   hm 20. oct. 2006 rev 1.5
    changed time_zone_offset from Real to INT, now in Minutes

   hm 27. feb. 2009 rev 1.6
    added type conversions to avoid warnings under codesys 3.0

   ks 13. nov. 2009 rev 1.7
    corrected error in formula

   *)
END_FUNCTION

FUNCTION "MINUTE" : Int   // FC197, SCL
TITLE = MINUTE
{ S7_Optimized_Access := 'FALSE' }
AUTHOR : hugo
FAMILY : TIDT
NAME : MINUTE
VERSION : 1.1
// extracts the minutes out of TOD truncating the ceconds
   VAR_INPUT
      itod : Time_Of_Day;
   END_VAR
BEGIN


     #MINUTE := DINT_TO_INT(T_CONV(#itod)/60000 - T_CONV(#itod)/3600000 * 60);


   (* change history

   2.10.2006 changes name of input to itod

   *)
END_FUNCTION

FUNCTION "MINUTE_OF_DT" : Int   // FC198, SCL
TITLE = MINUTE_OF_DT
{ S7_Optimized_Access := 'FALSE' }
AUTHOR : oscat
FAMILY : TIDT
NAME : M_DT
VERSION : 1.0
// MINUTE_OF_DT returns the current minute (minute of the hour) of a DT variable
   VAR_INPUT
      XDT : Date_And_Time;
      _XDT AT XDT : Array[0..7] of Byte;
   END_VAR
BEGIN


   #MINUTE_OF_DT := BCD16_TO_INT(#_XDT[4]); 

   (*
       original code:
       MINUTE_OF_DT := DWORD_TO_INT(DT_TO_DWORD(XDT) MOD 3600)/60;
   *)

   (* revision history
   hm      6.9.2008    rev 1.0
       original version


   *)
END_FUNCTION

FUNCTION "MINUTE_TO_TIME" : Time   // FC199, SCL
TITLE = MINUTE_TO_TIME
{ S7_Optimized_Access := 'FALSE' }
AUTHOR : hugo
FAMILY : TIDT
NAME : MIN2TI
VERSION : 1.2
// converts an amount of minutes in real to time
   VAR_INPUT
      IN : Real;
   END_VAR
BEGIN


   #MINUTE_TO_TIME := T_CONV(REAL_TO_DINT(#IN * 60000));


   (* revision history
   hm  4. aug 2006 rev 1.0
       original version

   hm  14. mar 2008    rev 1.1
       rounded the input after the last digit

   hm  24. feb. 2009   rev 1.2
       changed input to IN

   *)
END_FUNCTION

FUNCTION "MONTH_BEGIN" : Date   // FC200, SCL
TITLE = MONTH_BEGIN
{ S7_Optimized_Access := 'FALSE' }
AUTHOR : hugo
FAMILY : TIDT
NAME : MONBEG
VERSION : 1.0
// returns the date for the first day of the current month in the current year.
// 
// uses: DINT_DATE [FC404]
//       DATE_DINT [FC405]
//       DAY_OF_MONTH [FC178]
//       DAY_OF_YEAR [FC180] 
//       YEAR_BEGIN [FC217]
//       YEAR_OF_DATE [FC219]
//       LEAP_OF_DATE [FC193] 
//       LEAP_YEAR [FC194]
   VAR_INPUT
      idate : Date;
   END_VAR
BEGIN


   #MONTH_BEGIN := "DINT_DATE"("DATE_DINT"(#idate) - ("DAY_OF_MONTH"(#idate) - 1) * 86400);



   (* revision history
   hm  15. JUN: 2008   rev 1.0
       original version 


   *)
END_FUNCTION

FUNCTION "MONTH_END" : Date   // FC201, SCL
TITLE = MONTH_END
{ S7_Optimized_Access := 'FALSE' }
AUTHOR : hugo
FAMILY : TIDT
NAME : MONEND
VERSION : 1.1
// returns the date for the first day of the current month in the current year.
// 
// uses: DINT_DATE [FC404]
//       DATE_DINT [FC405]
//       SET_DATE [FC213]
//       LEAP_YEAR [FC194] 
//       YEAR_OF_DATE [FC219]
//       MONTH_OF_DATE [FC202]
//       DAY_OF_YEAR [FC180] 
//       YEAR_BEGIN [FC217]
//       LEAP_OF_DATE [FC193]
   VAR_INPUT
      idate : Date;
   END_VAR
BEGIN


   #MONTH_END := "DINT_DATE"("DATE_DINT"("SET_DATE"(YEAR:="YEAR_OF_DATE"(#idate),MONTH:="MONTH_OF_DATE"(#idate)+1,DAY:=1)) - 86400);

   (* revision history
   hm  15. jun. 2008   rev 1.0
       original version    

   hm  7. oct. 2008    rev 1.1
       changed function year to year_of_date
       changed function month to month_of_date

   *)
END_FUNCTION

FUNCTION "MONTH_OF_DATE" : Int   // FC202, SCL
TITLE = MONTH_OF_DATE
{ S7_Optimized_Access := 'FALSE' }
AUTHOR : hugo
FAMILY : TIDT
NAME : MONTH
VERSION : 1.3
// returns the month of a date  
// 
// uses: DAY_OF_YEAR [FC180]
//       YEAR_BEGIN [FC217] 
//       YEAR_OF_DATE [FC219] 
//       LEAP_OF_DATE [FC193]
//       LEAP_YEAR [FC194]
   VAR_INPUT
      IDATE : Date;
   END_VAR
BEGIN


   #MONTH_OF_DATE := "DAY_OF_YEAR"(#IDATE);
   IF #MONTH_OF_DATE < 32 THEN
       #MONTH_OF_DATE := 1;
   ELSIF "LEAP_OF_DATE"(#IDATE) THEN
       #MONTH_OF_DATE := (#MONTH_OF_DATE * 53 + 1668) / 1623;
   ELSE
       #MONTH_OF_DATE := (#MONTH_OF_DATE * 53 + 1700) / 1620;
   END_IF;


   (* code for rev 1.2
   MONTH_OF_DATE := DAY_OF_YEAR(IDATE);
   IF LEAP_OF_DATE(IDATE) THEN
       CASE MONTH_OF_DATE OF
           1..31   :   MONTH_OF_DATE := 1;
           32..60  :   MONTH_OF_DATE := 2;
           61..91  :   MONTH_OF_DATE := 3;
           92..121 :   MONTH_OF_DATE := 4;
           122..152:   MONTH_OF_DATE := 5;
           153..182:   MONTH_OF_DATE := 6;
           183..213:   MONTH_OF_DATE := 7;
           214..244:   MONTH_OF_DATE := 8;
           245..274:   MONTH_OF_DATE := 9;
           275..305:   MONTH_OF_DATE := 10;
           306..335:   MONTH_OF_DATE := 11;
           336..366:   MONTH_OF_DATE := 12;
       END_CASE;
   ELSE
       CASE MONTH_OF_DATE OF
           1..31   :   MONTH_OF_DATE := 1;
           32..59  :   MONTH_OF_DATE := 2;
           60..90  :   MONTH_OF_DATE := 3;
           91..120 :   MONTH_OF_DATE := 4;
           121..151:   MONTH_OF_DATE := 5;
           152..181:   MONTH_OF_DATE := 6;
           182..212:   MONTH_OF_DATE := 7;
           213..243:   MONTH_OF_DATE := 8;
           244..273:   MONTH_OF_DATE := 9;
           274..304:   MONTH_OF_DATE := 10;
           305..334:   MONTH_OF_DATE := 11;
           335..365:   MONTH_OF_DATE := 12;
       END_CASE;
   END_IF;
   *)


   (* revision history
   hm  1. aug 2006 rev 1.0
       original version    

   hm  1. okt 2007 rev 1.1
       replaced old code (string conversion) with mathematics
       the execution time is now multiple times faster.

   hm  7. oct. 2008    rev 1.2
       changed name of function from month to MONTH_OF_DATE

   hm  27. mar. 2009   rev 1.3
       new improved code

   *)
END_FUNCTION

FUNCTION "MULTIME" : Time   // FC203, SCL
TITLE = MULTIME
{ S7_Optimized_Access := 'FALSE' }
AUTHOR : hugo
FAMILY : TIDT
NAME : MULTIME
VERSION : 1.1
// multiplies a time by a real number and returns a time
   VAR_INPUT
      t : Time;
      "M" : Real;
   END_VAR
BEGIN


     #MULTIME := T_CONV(REAL_TO_DINT(DINT_TO_REAL(T_CONV(#t)) * #"M"));

   (* revision history
   hm      2. oct 2006 rev 1.0
       original version

   hm      14. mar 2008    rev 1.1
       rounded the result after the last digit

   *)
END_FUNCTION

FUNCTION "PERIOD" : Bool   // FC204, SCL
TITLE = PERIOD
{ S7_Optimized_Access := 'FALSE' }
AUTHOR : hugo
FAMILY : TIDT
NAME : PERIOD
VERSION : 1.3
// PERIOD checks if a given date is between two dates (d1 and d2) d1 is the starting date and d2 the last date for the period.
// the years of the dates are ignored, so the function period cheks for a time period within a year independet of the year.
// 
// uses: DAY_OF_YEAR [FC180]
//       YEAR_BEGIN [FC217] 
//       YEAR_OF_DATE [FC219] 
//       LEAP_OF_DATE [FC193]
//       LEAP_YEAR [FC194]
   VAR_INPUT
      d1 : Date;
      dx : Date;
      d2 : Date;
   END_VAR
   VAR_TEMP
      day1 : Int;
      day2 : Int;
      dayx : Int;
   END_VAR
BEGIN


   #day1 := "DAY_OF_YEAR"(#d1);
   #day2 := "DAY_OF_YEAR"(#d2);
   #dayx := "DAY_OF_YEAR"(#dx);
   IF NOT "LEAP_OF_DATE"(#dx) AND #dayx > 58 THEN #dayx := #dayx + 1; END_IF;
   IF NOT "LEAP_OF_DATE"(#d1) AND #day1 > 58 THEN #day1 := #day1 + 1; END_IF;
   IF NOT "LEAP_OF_DATE"(#d2) AND #day2 > 58 THEN #day2 := #day2 + 1; END_IF;

   IF #day2 < #day1 THEN
       (* the period spans over the new year *)
       #PERIOD := #dayx <= #day2 OR #dayx >= #day1;
   ELSE
       #PERIOD := #dayx >= #day1 AND #dayx <= #day2;
   END_IF;

   (* code before rev 1.2
   yx := year(dx);
   p1 := date_add(d1,0,0,0,yx - year(d1));
   p2 := date_add(d2,0,0,0,yx - year(d2));

   IF p2 >= p1 THEN
       period := dx <= p2  AND dx >= p1;
   ELSE
       period := dx <= p2 OR dx >= p1;
   END_IF;
   *)


   (* revision history

   hm      19. sep 2007    rev 1.0
       original version

   hm      20. sep 2007    rev 1.1
       corrected a problem with leap year

   hm      4. jan 2008     rev 1.2
       changed code for better performance

   hm      22. mar. 2008   rev 1.3
       function would deliver wrong results when d1, d2 or dx are a leap_year

   *)
END_FUNCTION

FUNCTION "PERIOD2" : Bool   // FC205, SCL
TITLE = PERIOD2
{ S7_Optimized_Access := 'FALSE' }
AUTHOR : hugo
FAMILY : TIDT
NAME : PERIOD2
VERSION : 1.0
// PERIOD2 checks if DX is within one of 4 periods and sets the output true if so.
   VAR_INPUT
      DP : Array[0..3, 0..1] of Date;
      DX : Date;
   END_VAR
BEGIN


   #PERIOD2 :=  (#DX >= #DP[0,0] AND #DX <= #DP[0,1]) OR
               (#DX >= #DP[1,0] AND #DX <= #DP[1,1]) OR
               (#DX >= #DP[2,0] AND #DX <= #DP[2,1]) OR
               (#DX >= #DP[3,0] AND #DX <= #DP[3,1]);


   (* revision history

   hm      27. apr 2008    rev 1.0
       original version


   *)
END_FUNCTION

FUNCTION "REFRACTION" : Real   // FC206, SCL
TITLE = REFRACTION
{ S7_Optimized_Access := 'FALSE' }
AUTHOR : hugo
FAMILY : TIDT
NAME : REFRACT
VERSION : 1.1
// REFRACTION calculates the atmospheric refraction in degrees.
// the input nangle goes from 0 at the hirizon to 90 at midday.
   VAR_INPUT
      ELEV : Real;
   END_VAR
   VAR_TEMP
      tmp : Real;
   END_VAR
BEGIN


   #tmp := LIMIT(MN:=-1.9, IN:=#ELEV, MX:=80.0);
   #REFRACTION := 0.0174532925199433 / TAN(0.0174532925199433 * (#tmp + 10.3 / (#tmp + 5.11)));


   (* revision histroy
   hm  14. jul. 2008   rev 1.0
       original release

   hm  7. mar. 2009    rev 1.1
       using new formula

   *)
END_FUNCTION

FUNCTION "SDT_TO_DATE" : Date   // FC207, SCL
TITLE = SDT_TO_DATE
{ S7_Optimized_Access := 'FALSE' }
AUTHOR : hugo
FAMILY : TIDT
NAME : SDT2DAT
VERSION : 1.0
// converts Structured date time (SDT) to Date Time
// 
// uses: SDT [UDT12]
//       SET_DATE [FC213]
//       LEAP_YEAR [FC194]
   VAR_INPUT
      DTI : "SDT";
   END_VAR
BEGIN


   #SDT_TO_DATE := "SET_DATE"(YEAR:=#DTI.YEAR,MONTH:=#DTI.MONTH,DAY:=#DTI.DAY);



   (* revision history

   hm 18. oct. 2008    rev 1.0
       original version

   *)
END_FUNCTION

FUNCTION "SDT_TO_DT" : Date_And_Time   // FC208, SCL
TITLE = SDT_TO_DT
{ S7_Optimized_Access := 'FALSE' }
AUTHOR : hugo
FAMILY : TIDT
NAME : SDT2DT
VERSION : 1.0
// converts Structured date time (SDT) to Date Time
// 
// uses: SDT [UDT12]
//       SET_DT [FC214]
   VAR_INPUT
      DTI : "SDT";
   END_VAR
   VAR_TEMP
      tSDT_TO_DT : Date_And_Time;
   END_VAR
BEGIN


   #tSDT_TO_DT := "SET_DT"(year:=#DTI.YEAR,month:=#DTI.MONTH,day:=#DTI.DAY,hour:=#DTI.HOUR,minute:=#DTI.MINUTE,second:=#DTI.SECOND);
   #SDT_TO_DT := #tSDT_TO_DT;

   (* revision history

   hm 18. oct. 2008    rev 1.0
       original version

   *)
END_FUNCTION

FUNCTION "SDT_TO_TOD" : Time_Of_Day   // FC209, SCL
TITLE = SDT_TO_TOD
{ S7_Optimized_Access := 'FALSE' }
AUTHOR : hugo
FAMILY : TIDT
NAME : SDT2TOD
VERSION : 1.1
// converts Structured date time (SDT) to Date Time
// 
// uses: SDT [UDT12]
   VAR_INPUT
      DTI : "SDT";
   END_VAR
BEGIN


   #SDT_TO_TOD := T_CONV(#DTI.HOUR * 3600000 + #DTI.MINUTE * 60000 + INT_TO_DINT(#DTI.SECOND) * 1000 + #DTI.MS);


   (* revision history

   hm 18. oct. 2008    rev 1.0
       original version

   hm  16. nov. 2008   rev 1.1
       added typecasts to avoid warnings
   *)
END_FUNCTION

FUNCTION "SECOND" : Real   // FC210, SCL
TITLE = SECOND
{ S7_Optimized_Access := 'FALSE' }
AUTHOR : hugo
FAMILY : TIDT
NAME : SEC
VERSION : 1.1
// returns the seconds and milliseconds as real of TOD
   VAR_INPUT
      itod : Time_Of_Day;
   END_VAR
BEGIN


     #SECOND := DINT_TO_REAL(T_CONV(#itod) - T_CONV(#itod)/60000 * 60000)/1000;



   (* change history

   2.10.2006 changes name of input to itod

   *)
END_FUNCTION

FUNCTION "SECOND_OF_DT" : Int   // FC211, SCL
TITLE = SECOND_OF_DT
{ S7_Optimized_Access := 'FALSE' }
AUTHOR : oscat
FAMILY : TIDT
NAME : S_DT
VERSION : 1.0
// SECOND_OF_DT returns the current second (second of minute) of a DT variable
   VAR_INPUT
      XDT : Date_And_Time;
      _XDT AT XDT : Array[0..7] of Byte;
   END_VAR
BEGIN


   #SECOND_OF_DT := BCD16_TO_INT(#_XDT[5]); 

   (*
       original code:
       SECOND_OF_DT := DWORD_TO_INT(DT_TO_DWORD(XDT) MOD 60);
   *)

   (* revision history
   hm      6.9.2008    rev 1.0
       original version


   *)
END_FUNCTION

FUNCTION "SECOND_TO_TIME" : Time   // FC212, SCL
TITLE = SECOND_TO_TIME
{ S7_Optimized_Access := 'FALSE' }
AUTHOR : hugo
FAMILY : TIDT
NAME : SEC2TI
VERSION : 1.2
// converts an amount of seconds in real to time
   VAR_INPUT
      IN : Real;
   END_VAR
BEGIN


   #SECOND_TO_TIME := T_CONV(REAL_TO_DINT(#IN * 1000));


   (* revision history
   hm  4. aug. 2006    rev 1.0
       original version

   hm  14. mar. 2008   rev 1.1
       rounded the input after the last digit

   hm  24. feb. 2009   rev 1.2
       changed input to IN
   *)
END_FUNCTION

FUNCTION "SET_DATE" : Date   // FC213, SCL
TITLE = SET_DATE
{ S7_Optimized_Access := 'FALSE' }
AUTHOR : hugo
FAMILY : TIDT
NAME : SETDATE
VERSION : 2.2
// creates a date output from year, month and day of month   
// 
// uses: LEAP_YEAR [FC194]
   VAR_INPUT
      YEAR : Int;
      MONTH : Int;
      DAY : Int;
   END_VAR
   VAR_TEMP
      count : DWord;
      MTH_OFS : Int;
   END_VAR
BEGIN


     (* only in Step 7 *)
     CASE LIMIT(MN:=1,IN:=#MONTH,MX:=12) OF
       1 : #MTH_OFS := 0;
       2 : #MTH_OFS := 31;
       3 : #MTH_OFS := 59;
       4 : #MTH_OFS := 90;
       5 : #MTH_OFS := 120;
       6 : #MTH_OFS := 151;
       7 : #MTH_OFS := 181;
       8 : #MTH_OFS := 212;
       9 : #MTH_OFS := 243;
       10 : #MTH_OFS := 273;
       11 : #MTH_OFS := 304;
       12 : #MTH_OFS := 334;
     ELSE:
       #MTH_OFS := 0;
     END_CASE;

     (* calculate the amount of days to 31.12. the year before *)
     #count := DINT_TO_DWORD(DWORD_TO_DINT(SHR(IN:=DINT_TO_DWORD(INT_TO_DINT(#YEAR) * 1461 - 2878172),N:=2)) + INT_TO_DINT(#DAY + #MTH_OFS));
     (* for leap years and month > february then add one more day *)
     IF #MONTH < 3 AND "LEAP_YEAR"(#YEAR) THEN
       #SET_DATE := T_CONV((DWORD_TO_DINT(#count) - 1) - 7305);
     ELSE
       #SET_DATE := T_CONV(DWORD_TO_DINT(#count) - 7305);
     END_IF;


   (*
   (* calculate the amount of days to 31.12. the year before *)
   count := DINT_TO_DWORD(DWORD_TO_DINT(SHR(IN:=DINT_TO_DWORD(INT_TO_DINT(year) * 1461 - 2878173),N:=2))+INT_TO_DINT(day));
   (* add the days for the month of the year *)
   CASE LIMIT(MN:=1,IN:=month,MX:=12) OF
       1 :           MTH_OFS := 0;
       2 :           MTH_OFS := 31;
       3 :           MTH_OFS := 59;
       4 :           MTH_OFS := 90;
       5 :           MTH_OFS := 120;
       6 :           MTH_OFS := 151;
       7 :           MTH_OFS := 181;
       8 :           MTH_OFS := 212;
       9 :           MTH_OFS := 243;
       10:           MTH_OFS := 273;
       11:           MTH_OFS := 304;
       12:           MTH_OFS := 334;
   ELSE: 
       MTH_OFS := 0;
   END_CASE ;

   count := DINT_TO_DWORD(DWORD_TO_DINT(count) + MTH_OFS);

   (* for leap years and month > february then add one more day *)
   IF month > 2 AND LEAP_YEAR(year) THEN count := DINT_TO_DWORD(DWORD_TO_DINT(count) + 1); END_IF;
   (* generate the date *)
   SET_DATE := DINT_TO_DATE(DWORD_TO_DINT(count) - 7305);


   (*
   count := DINT_TO_DWORD(DWORD_TO_DINT(SHR(IN:=DINT_TO_DWORD(INT_TO_DINT(year) * 1461 - 2878173),N:=2))+INT_TO_DINT(day));

   IF month < 5 THEN
       IF month < 3 THEN
           IF month = 2 THEN count := DINT_TO_DWORD(DWORD_TO_DINT(count) + 31); END_IF;
       ELSE
           IF month = 4 THEN
               count := DINT_TO_DWORD(DWORD_TO_DINT(count) + 90 + BOOL_TO_DINT(SHL(IN:=INT_TO_WORD(year),N:=14) = 0));
           ELSE (* month = 3 *)
               count := DINT_TO_DWORD(DWORD_TO_DINT(count) + 59 + BOOL_TO_DINT(SHL(IN:=INT_TO_WORD(year),N:=14) = 0));
           END_IF;
       END_IF;
   ELSIF month < 9 THEN
       IF month < 7 THEN
           IF month = 6 THEN
               count := DINT_TO_DWORD(DWORD_TO_DINT(count) + 151 + BOOL_TO_DINT(SHL(IN:=INT_TO_WORD(year),N:=14) = 0));
           ELSE (* month = 5 *)
               count := DINT_TO_DWORD(DWORD_TO_DINT(count) + 120 + BOOL_TO_DINT(SHL(IN:=INT_TO_WORD(year),N:=14) = 0));
           END_IF;
       ELSE
           IF month = 8 THEN
               count := DINT_TO_DWORD(DWORD_TO_DINT(count) + 212 + BOOL_TO_DINT(SHL(IN:=INT_TO_WORD(year),N:=14) = 0));
           ELSE (* month = 7 *)
               count := DINT_TO_DWORD(DWORD_TO_DINT(count) + 181 + BOOL_TO_DINT(SHL(IN:=INT_TO_WORD(year),N:=14) = 0));
           END_IF;
       END_IF;
   ELSE (* month is 9 or higher *)
       IF month < 11 THEN
           IF month = 10 THEN
               count := DINT_TO_DWORD(DWORD_TO_DINT(count) + 273 + BOOL_TO_DINT(SHL(IN:=INT_TO_WORD(year),N:=14) = 0));
           ELSE (* month = 9 *)
               count := DINT_TO_DWORD(DWORD_TO_DINT(count) + 243 + BOOL_TO_DINT(SHL(IN:=INT_TO_WORD(year),N:=14) = 0));
           END_IF;
       ELSE
           IF month = 12 THEN
               count := DINT_TO_DWORD(DWORD_TO_DINT(count) + 334 + BOOL_TO_DINT(SHL(IN:=INT_TO_WORD(year),N:=14) = 0));
           ELSE (* month = 11 *)
               count := DINT_TO_DWORD(DWORD_TO_DINT(count) + 304 + BOOL_TO_DINT(SHL(IN:=INT_TO_WORD(year),N:=14) = 0));
           END_IF;
       END_IF;
   END_IF;

   //SET_DATE := DWORD_TO_DATE(count * 86400);
   SET_DATE := DINT_TO_DATE(DWORD_TO_DINT(count) - 7305);
   *)



   (* revision history
   hm  4. aug. 2006    rev 1.0
       original version

   hm  19 sep. 2007    rev 1.1
       use function leap_year to calculate leap year, more exceptions are handled

   hm  1. okt  2007    rev 1.2
       added compatibility to step7

   hm  16.dec 2007     rev 1.3
       changed code to improove performance

   hm  3. jan. 2008    rev 1.4
       further improvements in performance

   hm  16. mar. 2008   rev 1.5
       added type conversions to avoid warnings under codesys 3.0

   hm  7. apr. 2008    rev 1.6
       deleted unused step7 code

   hm  14. oct. 2008   rev 1.7
       optimized code for better performance

   hm  25. oct. 2008   rev 2.0
       new code using setup constants
   *)*)


   (* revision history
   hm  4. aug. 2006  rev 1.0
     original version

   hm  19 sep. 2007  rev 1.1
     use function leap_year to calculate leap year, more exceptions are handled

   hm  1. okt  2007  rev 1.2
     added compatibility to step7

   hm  16.dec 2007   rev 1.3
     changed code to improove performance

   hm  3. jan. 2008  rev 1.4
     further improvements in performance

   hm  16. mar. 2008 rev 1.5
     added type conversions to avoid warnings under codesys 3.0

   hm  7. apr. 2008  rev 1.6
     deleted unused step7 code

   hm  14. oct. 2008 rev 1.7
     optimized code for better performance

   hm  25. oct. 2008 rev 2.0
     new code using setup constants

   hm  16. nov. 2008 rev 2.1
     added typecasts to avoid warnings

   hm  22. jan. 2011 rev 2.2
     improved performance
   *)
END_FUNCTION

FUNCTION "SET_DT" : Date_And_Time   // FC214, SCL
TITLE = SET_DT
{ S7_Optimized_Access := 'FALSE' }
AUTHOR : hugo
FAMILY : TIDT
NAME : SET_DT
VERSION : 1.5
// creates a date output from year, month and day of month
// year must be in the form of 4 digits ie 2006 or 1977.
   VAR_INPUT
      year : Int;
      month : Int;
      day : Int;
      hour : Int;
      minute : Int;
      second : Int;
   END_VAR
   VAR_TEMP
      tDT : Date_And_Time;
      _DT AT tDT : Array[0..7] of Byte;
      t_year : Int;
   END_VAR
BEGIN


     //set_DT := DWORD_TO_DT(DATE_TO_DWORD(set_Date(year, month, day)) + second + minute * 60 + INT_TO_DWORD(hour) * 3600);

     #t_year := #year - 1900;

     IF #t_year > 99 THEN 
       #t_year := #year - 2000; 
     END_IF;

     #_DT[0] := WORD_TO_BYTE(INT_TO_BCD16(#t_year));   // year
     #_DT[1] := WORD_TO_BYTE(INT_TO_BCD16(#month));    // month
     #_DT[2] := WORD_TO_BYTE(INT_TO_BCD16(#day));      // day
     #_DT[3] := WORD_TO_BYTE(INT_TO_BCD16(#hour));     // hour
     #_DT[4] := WORD_TO_BYTE(INT_TO_BCD16(#minute));   // minute
     #_DT[5] := WORD_TO_BYTE(INT_TO_BCD16(#second));   // second

     #SET_DT := #tDT;

   (* revision history
   hm  4. aug. 2006        rev 1.0
       original version

   hm      19 sep. 2007    rev 1.1
       use function leap_year to calculate leap year, more exceptions are handled

   hm      1. okt 2007     rev 1.2
       added step7 compatibility
       call function set_date

   hm      8. oct 2007     rev 1.3
       deleted unused variables count and leap

   hm      1. 11 2007      rev 1.4
       converted hour type integer to dword in calculation to avoid overrun on möller ecp4

   hm      16. mar 2008    rev 1.5
       added type conversions to avoid warnings under codesys 3.0
   *)
END_FUNCTION

FUNCTION "SET_TOD" : Time_Of_Day   // FC215, SCL
TITLE = SET_TOD
{ S7_Optimized_Access := 'FALSE' }
AUTHOR : hugo
FAMILY : TIDT
NAME : SET_TOD
VERSION : 1.5
// creates tod from hour minute and second
   VAR_INPUT
      hour : Int;
      minute : Int;
      second : Real;
   END_VAR
BEGIN


     #SET_TOD := T_CONV(REAL_TO_DINT(#second * 1000) + #minute * 60000 + #hour * 3600000);


   (* revision history

   hm      4.aug.2006      rev 1.0
       original version

   hm      11. sep 2007    rev 1.1
       changed coding to avoid a compiler warning under twincat.

   hm      1. nov 2007 rev 1.2
       changed coding to avoid possible overrun situation on möller ecp4

   hm      2. Nov  2007    rev 1.3
       changed dword to DINT in calcualtion to avoid warnings with some compilers

   hm      14. mar 2008    rev 1.4
       changed code to avoid rounding problem at last digit of millisecond

   hm      16. mar. 2008   rev 1.5
       added type conversions to avoid warning under codesys 3.0
   *)
END_FUNCTION

FUNCTION "WORK_WEEK" : Int   // FC216, SCL
TITLE = WORK_WEEK
{ S7_Optimized_Access := 'FALSE' }
AUTHOR : hugo
FAMILY : TIDT
NAME : WORKWE
VERSION : 1.5
// calculates the work week for a given date according to iso8601
// 
// uses: YEAR_OF_DATE [FC219]
//       YEAR_BEGIN [FC217]
//       DAY_OF_WEEK [FC179]
//       LEAP_YEAR [FC194]
   VAR_INPUT
      idate : Date;
   END_VAR
   VAR_TEMP
      d1 : Date;
      w1 : Int;
      ds : DInt;
      yr : Int;
      w31 : Int;
      w01 : Int;
      wm : Int;
   END_VAR
BEGIN


     (* berechne den 1.1 des jahres von idate. *)
     #yr := "YEAR_OF_DATE"(#idate);
     #d1 := "YEAR_BEGIN"(#yr);
     (* wochentag von d1 *)
     #w1 := "DAY_OF_WEEK"(#d1);
     (* offset des montags der eletzten KW des vorjahres *)
     (* wenn der erste tag des jahres größer als donnerstag ist dann beginnt die letzte kw am montag davor *)
     (* wenn der erste tag des jahres ein donnerstag oder kleiner ist beginnt die erste kw 2 montage davor *)
     IF #w1 < 5 THEN
       #ds := (T_CONV(#d1) + 7305) - (#w1 + 6);
     ELSE
       #ds := (T_CONV(#d1) + 7305) - (#w1 - 1);
     END_IF;

     (* kalenderwoche des eingangsdatums *)
     #WORK_WEEK := DINT_TO_INT(((T_CONV(#idate) + 7305) - #ds) / 7);

     (* korrektur wenn work_week = 0 *)
     IF #WORK_WEEK = 0 THEN
       (* work_week needs to be 53 when 1.jan of the year before is thursday or dec 31. is thursday. *)
       (* first and last weekday of a year is equal and one more day for a leap_year. *)
       IF #w1 > 1 THEN #w31 := #w1 - 1; ELSE #w31 := 7; END_IF;
       IF "LEAP_YEAR"(#yr - 1) AND #w31 > 1 THEN #w01 := #w31 - 1; ELSE #w1 := 7; END_IF;
       (* if first or last day of a year is a thursday, the year has 53 weeks *)
       #WORK_WEEK := 52 + BOOL_TO_INT(#w31 = 4 OR #w01 = 4);
     ELSE
       (* end of year calculation *)
       (* calculated the first and last weekday *)
       IF "LEAP_YEAR"(#yr) THEN
         IF #w1 < 7 THEN #w31 := #w1 + 1; ELSE #w31 := 1; END_IF;
       ELSE
         #w31 := #w1;
       END_IF;
       (* if first or last day is thursday then the year has 53 weeks otherwise only 52 *)
       #wm := 52 + BOOL_TO_INT(#w31 = 4 OR #w1 = 4);
       IF #WORK_WEEK > #wm THEN #WORK_WEEK := 1; END_IF;
     END_IF;



   (* old code before rev 1.2
   w1 := weekday(set_Date(year(idate), 1,1));
   IF w1 < 5 THEN
       work_week := (day_of_year(idate) + w1 + 5)/7;
   ELSE
       work_week := (day_of_year(idate) + w1 - 2)/7;
   END_IF
   *)


   (* revision history

   hm  17.1.2007       rev 1.1
       deleted unused variable yday

   hm  19. dec 2007    rev 1.2
       changed code for better performance
       changed code to comply with ISO8601

   hm  16. mar 2008    rev 1.3
       added type conversions to avoid warnings under codesys 3.0

   hm  7. oct. 2008    rev 1.4
       changed function year to year_of_date
       changed function weekday to day_of_week

   hm  25. oct. 2008   rev 1.5
       optimized code for performance
   *)
END_FUNCTION

FUNCTION "YEAR_BEGIN" : Date   // FC217, SCL
TITLE = YEAR_BEGIN
{ S7_Optimized_Access := 'FALSE' }
AUTHOR : hugo
FAMILY : TIDT
NAME : YEAR1ST
VERSION : 1.2
// returs the date of january 1st for the given year  
// the function works for dates from 1990 - 2100
   VAR_INPUT
      y : Int;
   END_VAR
BEGIN


   #YEAR_BEGIN := T_CONV(DWORD_TO_DINT(SHR(IN:=DINT_TO_DWORD(INT_TO_DINT(#y) * 1461 - 2878169),N:=2))-7305);

   (*
   year_begin := DWORD_TO_DATE(SHR(INT_TO_DWORD(y) * 1461 - 2878169,2)*86400);
   *)


   (* revision history
   hm  19. dec 2007    rev 1.0
       original version

   hm  4. jan 2008     rev 1.1
       formula for step7 was incorrect during leap years

   hm  7. apr. 2008    rev 1.2
       deleted unused step7 code
   *)
END_FUNCTION

FUNCTION "YEAR_END" : Date   // FC218, SCL
TITLE = YEAR_END
{ S7_Optimized_Access := 'FALSE' }
AUTHOR : hugo
FAMILY : TIDT
NAME : YEAREND
VERSION : 1.1
// returs the date of december 31st for the given year  
// the function works for dates from 1970 - 2099
   VAR_INPUT
      y : Int;
   END_VAR
BEGIN


     #YEAR_END := T_CONV(DWORD_TO_DINT(SHR(IN:=DINT_TO_DWORD(INT_TO_DINT(#y+1) * 1461 - 2878169),N:=2))-7305);
     // YEAR_END := DWORD_TO_DATE(SHR(INT_TO_DWORD(y) * 1461 - 2876712, 2) * 86400);


   (* revision history
   hm  15. jun. 2008 rev 1.0
     original version

   hm  24. jan 2011  rev 1.1
     improved performance
   *)

   (* revision history
   hm  15. jun. 2008 rev 1.0
     original version

   hm  24. jan 2011  rev 1.1
     improved performance
   *)
END_FUNCTION

FUNCTION "YEAR_OF_DATE" : Int   // FC219, SCL
TITLE = YEAR_OF_DATE
{ S7_Optimized_Access := 'FALSE' }
AUTHOR : hugo
FAMILY : TIDT
NAME : YEAR
VERSION : 1.4
// returs the year of a date  
// the function works for dates from 1990 - 2100
   VAR_INPUT
      IDATE : Date;
   END_VAR
BEGIN


   #YEAR_OF_DATE := DINT_TO_INT(((100 * T_CONV(#IDATE)) + 50) / 36525) + 1990;  

   (*
   year := DWORD_TO_INT((DATE_TO_DWORD(idate)+43200) / 31557600 + 1970);
   *)

   (* code used prior to rev 1.1
   year := DWORD_TO_INT((DATE_TO_DWORD(idate)/864+71954300)/36525);
   *)

   (* revision history
   hm  4. aug 2006     rev 1.0
       original version

   hm  1. okt 2007     rev 1.1
       corrected error in algorithm
       adjustment for S7 compatibility

   hm  23.12.2007      rev 1.2
       changed code for better performance

   hm  7. apr. 2008    rev 1.3
       deleted unused step7 code

   hm  7. oct. 2008    rev 1.4
       reneamed function (year) to year_of_date

   *)
END_FUNCTION

FUNCTION "DINT_DT" : Date_And_Time   // FC399, SCL
TITLE = DINT_DT
{ S7_Optimized_Access := 'FALSE' }
AUTHOR : dalbi
FAMILY : xS7
NAME : DINT_DT
VERSION : 1.0
// converts UNIX-Time to DATE_AND_TIME 
// max. 31.12.2089 23:59:59
// 
// uses: D_TOD_DT [FC3]
   VAR_INPUT
      IN : DInt;
   END_VAR
   VAR_TEMP
      CT : DInt;
      tIN : DInt;
      tIN1 : DInt;
      tIN2 : DInt;
      tDATI : Date_And_Time;
   END_VAR
BEGIN


     #tIN := #IN - 631152000; // correct DT 1. 1.1.1990 00:00:00

     // correct the Simatic DINT to UDINT
     IF #tIN < 0 THEN
         #tIN2 := #tIN + 2147483647;
         #tIN1 := 2147483647;
         #tIN2 := #tIN2 + 2;  // ?
       ELSE
         #tIN1 := #tIN;
         #tIN2 := 0;
     END_IF;

     #CT := TRUNC(DINT_TO_REAL(#tIN1) / 86400) + TRUNC(DINT_TO_REAL(#tIN2) / 86400); // calculate full days
     #tIN := (#tIN1 MOD 86400) + (#tIN2 MOD 86400); // calculate TOD in seconds

     #CT := #CT + TRUNC(DINT_TO_REAL(#tIN) / 86400);
     #tIN := #tIN MOD 86400;

     #tDATI := T_COMBINE(IN1:=T_CONV(#CT),IN2:=T_CONV(#tIN * 1000));
     #DINT_DT := #tDATI;
END_FUNCTION

FUNCTION "DT_DINT" : DInt   // FC400, SCL
TITLE = DT_DINT
{ S7_Optimized_Access := 'FALSE' }
AUTHOR : dalbi
FAMILY : xS7
NAME : DT_DINT
VERSION : 1.0
// converts DATE_AND_TIME to UNIX-Time max. 31.12.2089 23:59:59
// 
// uses: DT_DATE [FC6]
//       DT_TOD [FC8]
   VAR_INPUT
      DATI : Date_And_Time;
   END_VAR
   VAR_TEMP
      tDATI : Date_And_Time;
   END_VAR
BEGIN


     #tDATI := #DATI;
     #DT_DINT := (T_CONV(T_CONV(#tDATI)) + 7305) * 86400;  
     #DT_DINT := #DT_DINT + T_CONV(T_CONV(#tDATI)) / 1000;
END_FUNCTION

FUNCTION "UTC_TO_LTIME" : Date_And_Time   // FC402, SCL
TITLE = UTC_TO_LTIME
{ S7_Optimized_Access := 'FALSE' }
AUTHOR : oscat
FAMILY : TIDT
NAME : LTIME
VERSION : 1.9
// ltime is a real time clock that uses the system rtc as utc time and calculates and given time zone.
// the utc time is supplied on the input UTC.
// according to the input variable time_zone_offset when the input dst_enable is true,
// the dst on and off times are calculated by a formula for any given year and the time is advanced and reset by one hour
// at 02:00 and 03:00 for the last sunday of march and last sunday of october.
// the code is high performance and the rtc counts every second.
// if more then one time zone is needed by the systen the clock can be started many times by placing more then one function block.
// 
// uses: DST [FC183]
//       YEAR_OF_DATE [FC219] 
//       DT_DATE [FC6] 
//       DT_DINT [FC400] 
//       DT_TOD [FC8]
//       SET_DT [FC214] 
//       DINT_DT [FC399]
//       D_TOD_DT [FC3]
   VAR_INPUT
      UTC : Date_And_Time;
      DST_ENABLE : Bool;
      TIME_ZONE_OFFSET : Int;
   END_VAR
   VAR_TEMP
      tmp : Int;
      tUTC : Date_And_Time;
      tLTIME : Date_And_Time;
   END_VAR
BEGIN


   #tUTC := #UTC;
   #tLTIME := #UTC_TO_LTIME;

   #tmp := #TIME_ZONE_OFFSET * 60 + BOOL_TO_INT(#DST_ENABLE AND "DST"(#tUTC)) * 3600;
   IF #tmp < 0 THEN
       #tmp := ABS(#tmp);
       #tLTIME := "DINT_DT"("DT_DINT"(#tUTC) -  INT_TO_DINT(#tmp));
   ELSE
       #tLTIME := "DINT_DT"("DT_DINT"(#tUTC) +  INT_TO_DINT(#tmp));
   END_IF;

   #UTC_TO_LTIME := #tLTIME;

   (* revision history

   hm 2.10.2006    rev 1.1
       corrected an error where dst would be delayed by 0.1second

   hm 17.1.2007    rev 1.2
       added utc input instead of internal sysrtcgettime because this would only work on wago.
       dst_enable would not be checked before dst would be enabled.

   hm 18.3.2007    rev 1.3
       changed code, dst would not work during first cycle.

   hm 24.10.2007   rev 1.4
       changed code because the execution every 100ms can cause major problems if the supplied time was not correct at start.
       use of new dst function

   hm 12. nov 2007 rev 1.5
           changed Type of time_zone_offset from time to int to allow for time zones with negative offset

   hm  8 dec 2007      rev 1.6
       corrected a problem with time_zone_offset

   hm  14. oct. 2008   rev 1.7
       renamed module from LTIME to UTC_TO_LTIME
       changed function weekday to day_of_week
       optimized code for better performance

   hm  20. oct. 2008   rev 1.8
       changes type of input TIME_ZONE_OFFSET from real to int, now is in +/-minutes
       deleted outputs DST_ON and WDAY
       converted to function

   hm  27. feb. 2009   rev 1.9
       added type conversions to avoid warnings under codesys 3.0

   *)
END_FUNCTION

FUNCTION "DINT_DATE" : Date   // FC404, SCL
TITLE = DINT_DATE
{ S7_Optimized_Access := 'FALSE' }
AUTHOR : dalbi
FAMILY : xS7
NAME : DINT_D
VERSION : 1.0
// convert IEC-DATE to S7 DATE
   VAR_INPUT
      D : DInt;
   END_VAR
   VAR_TEMP
      temp_D : DInt;
      _temp_D AT temp_D : Array[0..31] of Bool;
   END_VAR
BEGIN


     #temp_D := #D - 631152000;

     IF #temp_D < 0 THEN
       #_temp_D[7] := FALSE;
       #temp_D := TRUNC(DINT_TO_REAL(#temp_D) / 86400) + 24856;
     ELSE
       #temp_D := #temp_D / 86400;
     END_IF;

     #DINT_DATE := T_CONV(#temp_D);
END_FUNCTION

FUNCTION "DATE_DINT" : DInt   // FC405, SCL
TITLE = DATE_DINT
{ S7_Optimized_Access := 'FALSE' }
AUTHOR : dalbi
FAMILY : xS7
NAME : D_DINT
VERSION : 1.0
// convert S7 DATE to IEC-DATE
   VAR_INPUT
      D : Date;
   END_VAR
BEGIN


   (* 1.1.1990 00:00:00 = 631152000 *)
   #DATE_DINT := T_CONV(#D) * 86400 + 631152000;
END_FUNCTION

FUNCTION "DAYS_IN_MONTH" : Int   // FC415, SCL
TITLE = DAYS_IN_MONTH
{ S7_Optimized_Access := 'FALSE' }
AUTHOR : hugo
FAMILY : TIDT
NAME : DAYiMON
VERSION : 1.0
// returs the total days of the current month. e.g. 31 for january.
// the function works for dates from 1990 - 2168
// 
// uses: DAY_OF_YEAR [FC180]
//       YEAR_BEGIN [FC217] 
//       YEAR_OF_DATE [FC219] 
//       LEAP_OF_DATE [FC193]
//       LEAP_YEAR [FC194]
   VAR_INPUT
      IDATE : Date;
   END_VAR
BEGIN


   #DAYS_IN_MONTH := "DAY_OF_YEAR"(#IDATE);
   IF "LEAP_OF_DATE"(#IDATE) THEN
       CASE #DAYS_IN_MONTH OF
           32..60  :   #DAYS_IN_MONTH := 29;
           92..121 :   #DAYS_IN_MONTH := 30;
           153..182:   #DAYS_IN_MONTH := 30;
           245..274:   #DAYS_IN_MONTH := 30;
           306..335:   #DAYS_IN_MONTH := 30;
       ELSE
           #DAYS_IN_MONTH := 31;
       END_CASE;
   ELSE
       CASE #DAYS_IN_MONTH OF
           32..59  :   #DAYS_IN_MONTH := 28;
           91..120 :   #DAYS_IN_MONTH := 30;
           152..181:   #DAYS_IN_MONTH := 30;
           244..273:   #DAYS_IN_MONTH := 30;
           305..334:   #DAYS_IN_MONTH := 30;
       ELSE
           #DAYS_IN_MONTH := 31;
       END_CASE;
   END_IF;



   (* revision history
   hm  27. mar. 2009       rev 1.0
       original version

   *)
END_FUNCTION

FUNCTION "DAYS_IN_YEAR" : Int   // FC416, SCL
TITLE = DAYS_IN_YEAR
{ S7_Optimized_Access := 'FALSE' }
AUTHOR : hugo
FAMILY : TIDT
NAME : DAYiYEAR
VERSION : 1.0
// returs the total days of the year.
// the function retruns 366 for leap years and 365 otherwise.
// the function works for dates from 1970 - 2099
// 
// uses: LEAP_OF_DATE [FC193]
//       LEAP_YEAR [FC194] 
//       YEAR_OF_DATE [FC219]
   VAR_INPUT
      IDATE : Date;
   END_VAR
BEGIN


   IF "LEAP_OF_DATE"(#IDATE) THEN
       #DAYS_IN_YEAR := 366;
   ELSE
       #DAYS_IN_YEAR := 365;
   END_IF;


   (* revision history
   hm  27. mar. 2009       rev 1.0
       original version

   *)
END_FUNCTION

FUNCTION "TIMECHECK" : Bool   // FC418, SCL
TITLE = TIMECHECK
{ S7_Optimized_Access := 'FALSE' }
AUTHOR : oscat
FAMILY : TIDT
NAME : TIMCHK
VERSION : 1.0
// this function retruns true if the daytime TD is between start and stop and returns true if so.
// if you want to generate an event to span over midnight, start timemust be later than the stop time.
   VAR_INPUT
      TD : Time_Of_Day;
      START : Time_Of_Day;
      STOP : Time_Of_Day;
   END_VAR
BEGIN


   IF #STOP < #START THEN
     #TIMECHECK := #START <= #TD OR #TD < #STOP;
   ELSE
     #TIMECHECK := #START <= #TD AND #TD < #STOP;
   END_IF;


   (* revision history
   hm 19. jul. 2009  rev 1.0
     original release

   *)
END_FUNCTION

FUNCTION "SUN_MIDDAY" : Time_Of_Day   // FC432, SCL
TITLE = SUN_MIDDAY
{ S7_Optimized_Access := 'FALSE' }
AUTHOR : hugo
FAMILY : TIDT
NAME : SUNMID
VERSION : 1.0
// this FUNCTION calculates the time when the sun stand exactly south of a given location.
// 
// uses:  DAY_OF_YEAR (FC180)
//        DATE_DINT (FC405)
//        HOUR_TO_TOD (FC190)
   VAR_INPUT
      LON : Real;
      UTC : Date;
   END_VAR
   VAR_TEMP
      T : Real;
      OFFSET : Real;
   END_VAR
BEGIN


   #T := INT_TO_REAL("DAY_OF_YEAR"(#UTC));
   #OFFSET := -0.1752 * SIN(0.033430 * #T + 0.5474) - 0.1340 * SIN(0.018234 * #T - 0.1939);
   #SUN_MIDDAY := "HOUR_TO_TOD"(12.0 - #OFFSET - #LON * 0.0666666666666);


   (* revision history

   hm  26. jan. 2011 rev 1.0
     initial release

   *)
END_FUNCTION

// ===== PLC "xS7"  Unspecific CPU S7 300 =====

DATA_BLOCK "TEMP"   // DB7
TITLE = temporary Strings
{ S7_Optimized_Access := 'FALSE' }
AUTHOR : dalbi
FAMILY : xS7
NAME : DBTEMP
VERSION : 1.1
   VAR
      STR1 : String[254];
      STR2 : String[254];
      STR3 : String[254];
      TEMP : String[254];
   END_VAR
BEGIN
END_DATA_BLOCK

DATA_BLOCK "IDB_STIME"   // DB64
{ S7_Optimized_Access := 'FALSE' }
AUTHOR : dalbi
FAMILY : MEASURE
VERSION : 0.0
// stored: InstanceOfName STIME
"STIME"
BEGIN
END_DATA_BLOCK

FUNCTION_BLOCK "STIME"   // FB64, SCL
TITLE = STIME
{ S7_Optimized_Access := 'FALSE' }
AUTHOR : dalbi
FAMILY : MEASURE
NAME : STIME
VERSION : 1.4
// this function block makes sure that the timer of a siemens sps counts from 0 - 2^32-1.
   VAR_OUTPUT
      tx : DWord;
      at_tx AT tx : Array[0..31] of Bool;
   END_VAR
   VAR
      last_time : DWord;
      bit31 : Bool;
      init : Bool := TRUE;
   END_VAR
   VAR_TEMP
      TOP_SI : Struct
         EV_CLASS : Byte;
         EV_NUM : Byte;
         PRIORITY : Byte;
         NUM : Byte;
         TYP2_3 : Byte;
         TYP1 : Byte;
         ZI1 : Word;
         ZI2_3 : DWord;
      END_STRUCT;
      START_UP_SI : Struct
         EV_CLASS : Byte;
         EV_NUM : Byte;
         PRIORITY : Byte;
         NUM : Byte;
         TYP2_3 : Byte;
         TYP1 : Byte;
         ZI1 : Word;
         ZI2_3 : DWord;
      END_STRUCT;
      ERR : Int;
   END_VAR
BEGIN


   (* this FB is only necessary for siemens sps
   the siemens sps timer counts from 0 to 2^31-1 and starts at 0 sfter overrun.
   this means that the bit 31 (the highest bit ) will never be used and therefore
   a problem arises when t2 - t1 is checked.
   t2 - t1 is always valid also in an timer overrun situation where the time t1 is very high and t2 is very low.
   the result of the subtraction t2 - t1 however is still valid.
   this calculation does not work for soiemens because the highest bit is not used.

   this module stores the highest bit, changes the highest bit at every overrun occurence and stuffs ther highest bit in the output.
   the output is then used by t_plc_us and t_plc_ms.

   the correction needs and fb and not a function because the value of the highest bit has to be stored.

   do never use this function block in a codesys environment. the timer in codesys is correct and runs from 0 to 2^32-1
   *)

   (* read actual startup info *)
   (* OB1_SCAN_1  BYTE  -  B#16#01: Abschluss des Neustarts (Warmstarts)
                        -  B#16#02: Abschluss des Wiederanlaufs
                        -  B#16#03: Abschluss des freien Zyklus
                        -  B#16#04: Abschluss des Kaltstarts
                        -  B#16#05: Erster OB 1-Zyklus der neuen Master-CPU nach 
                                    Master-Reserve-Umschaltung und STOP des 
                                    bisherigen Masters *)

   #ERR := RD_SINFO (TOP_SI => #TOP_SI, START_UP_SI => #START_UP_SI);

   (* reset last_time on system startup *)
   IF #TOP_SI.EV_NUM = 1 OR #TOP_SI.EV_NUM = 2 OR #TOP_SI.EV_NUM = 4 OR NOT #init THEN 
       #last_time := 0;
       #bit31 := false;
       #init := true;
   END_IF;

   (* read the system timer *)
   #tx := DINT_TO_DWORD(T_CONV(TIME_TCK()));

   (* check for overrun *)
   IF DWORD_TO_DINT(#tx) < DWORD_TO_DINT(#last_time) THEN
       (* an overrun has occured, change the value of the highest bit *)
       #bit31 := NOT #bit31;
   END_IF;

   (* stuff the highest bit into the timer value *)
   #at_tx[7] := #bit31;

   (* remember the last system time for the next overrun check *)
   #last_time := #tx;


   (* revision history
   DA  14.9.2007 rev 1.0
     original version

   DA  24.2.2008 rev 1.1
     added self reset on system startup

   DA   2.5.2008 rev 1.2
     corect a problem running under OB35

   DA  12.3.2009 rev 1.3
     corect a problem run on different CPUs

   DA  22.12.2009 rev 1.4
     corect a problem on startup
   *)
END_FUNCTION_BLOCK

FUNCTION_BLOCK "R_TRIG"   // FB235, SCL
TITLE = R_TRIG
{ S7_Optimized_Access := 'FALSE' }
AUTHOR : dalbi
FAMILY : xS7
NAME : R_TRIG
VERSION : 1.0
// detect rising edge
   VAR_INPUT
      CLK : Bool;
   END_VAR
   VAR_OUTPUT
      Q : Bool;
   END_VAR
   VAR
      "M" : Bool;
   END_VAR
BEGIN


     #Q := #CLK AND NOT #"M";
     #"M" := #CLK;
END_FUNCTION_BLOCK

FUNCTION_BLOCK "F_TRIG"   // FB236, SCL
TITLE = F_TRIG
{ S7_Optimized_Access := 'FALSE' }
AUTHOR : dalbi
FAMILY : xS7
NAME : F_TRIG
VERSION : 1.0
// detect falling edge
   VAR_INPUT
      CLK : Bool;
   END_VAR
   VAR_OUTPUT
      Q : Bool;
   END_VAR
   VAR
      "M" : Bool;
   END_VAR
BEGIN


    #Q := NOT #CLK AND #"M";
    #"M" := #CLK;
END_FUNCTION_BLOCK

FUNCTION "DINT_DT" : Date_And_Time   // FC399, SCL
TITLE = DINT_DT
{ S7_Optimized_Access := 'FALSE' }
AUTHOR : dalbi
FAMILY : xS7
NAME : DINT_DT
VERSION : 1.0
// converts UNIX-Time to DATE_AND_TIME 
// max. 31.12.2089 23:59:59
// 
// uses: D_TOD_DT [FC3]
   VAR_INPUT
      IN : DInt;
   END_VAR
   VAR_TEMP
      CT : DInt;
      tIN : DInt;
      tIN1 : DInt;
      tIN2 : DInt;
      tDATI : Date_And_Time;
   END_VAR
BEGIN


     #tIN := #IN - 631152000; // correct DT 1. 1.1.1990 00:00:00

     // correct the Simatic DINT to UDINT
     IF #tIN < 0 THEN
         #tIN2 := #tIN + 2147483647;
         #tIN1 := 2147483647;
         #tIN2 := #tIN2 + 2;  // ?
       ELSE
         #tIN1 := #tIN;
         #tIN2 := 0;
     END_IF;

     #CT := TRUNC(DINT_TO_REAL(#tIN1) / 86400) + TRUNC(DINT_TO_REAL(#tIN2) / 86400); // calculate full days
     #tIN := (#tIN1 MOD 86400) + (#tIN2 MOD 86400); // calculate TOD in seconds

     #CT := #CT + TRUNC(DINT_TO_REAL(#tIN) / 86400);
     #tIN := #tIN MOD 86400;

     #tDATI := T_COMBINE(IN1:=T_CONV(#CT),IN2:=T_CONV(#tIN * 1000));
     #DINT_DT := #tDATI;
END_FUNCTION

FUNCTION "DT_DINT" : DInt   // FC400, SCL
TITLE = DT_DINT
{ S7_Optimized_Access := 'FALSE' }
AUTHOR : dalbi
FAMILY : xS7
NAME : DT_DINT
VERSION : 1.0
// converts DATE_AND_TIME to UNIX-Time max. 31.12.2089 23:59:59
// 
// uses: DT_DATE [FC6]
//       DT_TOD [FC8]
   VAR_INPUT
      DATI : Date_And_Time;
   END_VAR
   VAR_TEMP
      tDATI : Date_And_Time;
   END_VAR
BEGIN


     #tDATI := #DATI;
     #DT_DINT := (T_CONV(T_CONV(#tDATI)) + 7305) * 86400;  
     #DT_DINT := #DT_DINT + T_CONV(T_CONV(#tDATI)) / 1000;
END_FUNCTION

FUNCTION "EQ_ANY" : Bool   // FC401, SCL
TITLE = EQ_ANY
{ S7_Optimized_Access := 'FALSE' }
AUTHOR : dalbi
FAMILY : xS7
NAME : EQ_ANY
VERSION : 1.0
   VAR_INPUT
      IN1 : ANY;
      IN2 : ANY;
   END_VAR
   VAR_TEMP
      tANY1 : ANY;
      _ANY1 AT tANY1 : Struct
         id : Byte;
         DataType : Byte;
         Lenght : Word;
         DBNr : Word;
         Byte_Pointer : DWord;
      END_STRUCT;
      tANY2 : ANY;
      _ANY2 AT tANY2 : Struct
         id : Byte;
         DataType : Byte;
         Lenght : Word;
         DBNr : Word;
         Byte_Pointer : DWord;
      END_STRUCT;
      tAdr1 : Int;
      tAdr2 : Int;
      i : Int;
   END_VAR
BEGIN


     #tANY1 := #IN1;
     #tANY2 := #IN2;

     #tAdr1 := DWORD_TO_INT(SHR(IN:=SHL(IN:=#_ANY1.Byte_Pointer,N:=8),N:=11));
     #tAdr2 := DWORD_TO_INT(SHR(IN:=SHL(IN:=#_ANY2.Byte_Pointer,N:=8),N:=11));

     #EQ_ANY := TRUE;

     IF #_ANY1.Lenght <> #_ANY2.Lenght THEN
       #EQ_ANY := FALSE;
     ELSE
       FOR #i := 0 TO WORD_TO_INT(#_ANY1.Lenght)-1 DO
         IF WORD_TO_BLOCK_DB(#_ANY1.DBNr).DB(#tAdr1+#i) <> WORD_TO_BLOCK_DB(#_ANY2.DBNr).DB(#tAdr2+#i) THEN
           #EQ_ANY := FALSE;
           EXIT;
         END_IF;
       END_FOR;
     END_IF;
END_FUNCTION

FUNCTION "DINT_DATE" : Date   // FC404, SCL
TITLE = DINT_DATE
{ S7_Optimized_Access := 'FALSE' }
AUTHOR : dalbi
FAMILY : xS7
NAME : DINT_D
VERSION : 1.0
// convert IEC-DATE to S7 DATE
   VAR_INPUT
      D : DInt;
   END_VAR
   VAR_TEMP
      temp_D : DInt;
      _temp_D AT temp_D : Array[0..31] of Bool;
   END_VAR
BEGIN


     #temp_D := #D - 631152000;

     IF #temp_D < 0 THEN
       #_temp_D[7] := FALSE;
       #temp_D := TRUNC(DINT_TO_REAL(#temp_D) / 86400) + 24856;
     ELSE
       #temp_D := #temp_D / 86400;
     END_IF;

     #DINT_DATE := T_CONV(#temp_D);
END_FUNCTION

FUNCTION "DATE_DINT" : DInt   // FC405, SCL
TITLE = DATE_DINT
{ S7_Optimized_Access := 'FALSE' }
AUTHOR : dalbi
FAMILY : xS7
NAME : D_DINT
VERSION : 1.0
// convert S7 DATE to IEC-DATE
   VAR_INPUT
      D : Date;
   END_VAR
BEGIN


   (* 1.1.1990 00:00:00 = 631152000 *)
   #DATE_DINT := T_CONV(#D) * 86400 + 631152000;
END_FUNCTION

FUNCTION "SYS_STARTUP" : Byte   // FC407, SCL
TITLE = System Startup
{ S7_Optimized_Access := 'FALSE' }
AUTHOR : dalbi
FAMILY : xS7
NAME : SYSON
VERSION : 1.0
// detect system startup
   VAR_IN_OUT
      Startup : Bool;
   END_VAR
   VAR_TEMP
      TOP_SI : Struct
         EV_CLASS : Byte;
         EV_NUM : Byte;
         PRIORITY : Byte;
         NUM : Byte;
         TYP2_3 : Byte;
         TYP1 : Byte;
         ZI1 : Word;
         ZI2_3 : DWord;
      END_STRUCT;
      START_UP_SI : Struct
         EV_CLASS : Byte;
         EV_NUM : Byte;
         PRIORITY : Byte;
         NUM : Byte;
         TYP2_3 : Byte;
         TYP1 : Byte;
         ZI1 : Word;
         ZI2_3 : DWord;
      END_STRUCT;
      ERR : Int;
   END_VAR
BEGIN


   (* read actual startup info *)
   (* OB1_SCAN_1  BYTE  -  B#16#01: Abschluss des Neustarts (Warmstarts)
                        -  B#16#02: Abschluss des Wiederanlaufs
                        -  B#16#03: Abschluss des freien Zyklus
                        -  B#16#04: Abschluss des Kaltstarts
                        -  B#16#05: Erster OB 1-Zyklus der neuen Master-CPU nach 
                                    Master-Reserve-Umschaltung und STOP des 
                                    bisherigen Masters *)

     #ERR := RD_SINFO (TOP_SI => #TOP_SI, START_UP_SI => #START_UP_SI);

   (* detect system startup *)
     IF #TOP_SI.EV_NUM <> 3 THEN 
       #Startup := TRUE;
     END_IF;  

     #SYS_STARTUP := #TOP_SI.EV_NUM;
END_FUNCTION

FUNCTION "EXPT" : Real   // FC408, SCL
TITLE = EXPT
{ S7_Optimized_Access := 'FALSE' }
AUTHOR : dalbi
FAMILY : xS7
NAME : EXPT
VERSION : 1.0
// potentialization of variable with other
   VAR_INPUT
      X : Real;
      N : Real;
   END_VAR
BEGIN


     #EXPT := #X ** #N;
END_FUNCTION

FUNCTION "BYTE_TO_STRING" : String[254]   // FC417, SCL
TITLE = BYTE_TO_STRING
{ S7_Optimized_Access := 'FALSE' }
AUTHOR : dalbi
FAMILY : xS7
NAME : BY2STR
VERSION : 1.0
// convert BYTE(USINT) to STRING[3]
   VAR_INPUT
      "B" : Byte;
   END_VAR
   VAR_TEMP
      bw : Word;
      str : Struct
         Maximal : Byte;
         Actual : Byte;
         CHR : Array[1..3] of Byte;
      END_STRUCT;
      tSTR AT str : String [ 3 ];   // MigChange: STRING[3]
   END_VAR
BEGIN


   (* tSTR initialisieren *)
   #str.Maximal := 3;

   (* BYTE in BCD wandeln *)
   #bw := INT_TO_BCD16(BYTE_TO_INT(#"B"));

   (* STRING erstellen *)
   IF BCD16_TO_INT(#bw) > 99 THEN     //BCD von 99..255
       #str.Actual := 3;
       #str.CHR[1] := WORD_TO_BYTE(SHR(IN:=#bw AND W#16#0F00, N:=8) OR 16#30);
       #str.CHR[2] := WORD_TO_BYTE(SHR(IN:=#bw AND W#16#00F0, N:=4) OR 16#30);
       #str.CHR[3] := WORD_TO_BYTE(#bw AND W#16#000F OR 16#30);
   ELSIF BCD16_TO_INT(#bw) > 9 THEN   //BCD von 10..99
       #str.Actual := 2;
       #str.CHR[1] := WORD_TO_BYTE(SHR(IN:=#bw AND W#16#00F0, N:=4) OR 16#30);
       #str.CHR[2] := WORD_TO_BYTE(#bw AND W#16#000F OR 16#30);
   ELSE                            //BCD von 0..9
       #str.Actual := 1;
       #str.CHR[1] := WORD_TO_BYTE(#bw AND W#16#000F OR 16#30);
   END_IF;

   (* Temporären STRING nach OUT kopieren *)
   #BYTE_TO_STRING := #tSTR;


   (* revision history

   da 10.04.2009       rev 1.0

   *)
END_FUNCTION